
screen "St_Output Bundled_1" 320x240
   IOField "I/O field_9" at 228,67 size 87x20; FormatPattern 999.99
      ProcessValue <- "Data_Real_% label Sloft[1]"
   IOField "I/O field_10" at 228,86 size 87x20; FormatPattern 999.99
      ProcessValue <- "Data_Real_% Unlabel Sloft[1]"
   TextField "Text field_1" at 4,0 size 268x18; Text 'CURRENT SHIFT MINUS 1 ( Output Bundle )'
   IOField "I/O field_2" at 145,86 size 84x20; FormatPattern 9999999
      ProcessValue <- "Data_IntData_Un label Sloft[1]"
   IOField "I/O field_3" at 145,67 size 84x20; FormatPattern 9999999
      ProcessValue <- "Data_IntData_Label Sloft[1]"
   IOField "I/O field_6" at 6,17 size 109x15; FormatPattern 9999999999999999999999999999999999999999
      ProcessValue <- "Data_DTL1_Cur_ShiftA_1"
   TextField "Text field_9" at 120,17 size 18x13; Text 'S/D'
   IOField "I/O field_7" at 143,17 size 109x15; FormatPattern 9999999999999999999999999999999999999999
      ProcessValue <- "Data_DTL1_Cur_ShiftB_1"
   Button "Button_1" at 101,214 size 128x25; TextOff 'Back To Quantity Data'; TextOn 'Page 1'
      on Click: ActivateScreen("St_Quantity Data_1", 0)
   TextField "Text field_5" at 7,86 size 139x20; Text 'Unlabeled Bundle'
   TextField "Text field_4" at 7,67 size 139x20; Text 'Labeled Bundle'
   TextField "Text field_15" at 145,48 size 84x19; Text 'Pcs'
   TextField "Text field_16" at 228,48 size 87x19; Text '% (From input)'
   TextField "Text field_17" at 7,48 size 139x19; Text 'Output Bundle'
   IOField "I/O field_27" at 253,16 size 66x17; FormatPattern ????????
      ProcessValue <- "Data_String_sDT_Machine id"

screen "St_Output Bundled_2" 320x240
   IOField "I/O field_9" at 228,67 size 87x20; FormatPattern 999.99
      ProcessValue <- "Data_Real_% label Sloft[2]"
   IOField "I/O field_10" at 228,86 size 87x20; FormatPattern 999.99
      ProcessValue <- "Data_Real_% Unlabel Sloft[2]"
   TextField "Text field_1" at 4,0 size 262x18; Text 'CURRENT SHIFT MINUS 2 ( Ouput Bundle )'
   IOField "I/O field_2" at 145,86 size 84x20; FormatPattern 9999999
      ProcessValue <- "Data_IntData_Un label Sloft[2]"
   IOField "I/O field_3" at 145,67 size 84x20; FormatPattern 9999999
      ProcessValue <- "Data_IntData_Label Sloft[2]"
   IOField "I/O field_6" at 6,17 size 109x15; FormatPattern 9999999999999999999999999999999999999999
      ProcessValue <- "Data_DTL1_Cur_ShiftA_2"
   TextField "Text field_9" at 120,17 size 18x13; Text 'S/D'
   IOField "I/O field_7" at 143,17 size 109x15; FormatPattern 9999999999999999999999999999999999999999
      ProcessValue <- "Data_DTL1_Cur_ShiftB_2"
   Button "Button_1" at 101,214 size 128x25; TextOff 'Back To Quantity Data'; TextOn 'Page 1'
      on Click: ActivateScreen("St_Quantity Data_2", 0)
   TextField "Text field_5" at 7,86 size 139x20; Text 'Unlabeled Bundle'
   TextField "Text field_4" at 7,67 size 139x20; Text 'Labeled Bundle'
   TextField "Text field_15" at 145,48 size 84x19; Text 'Pcs'
   TextField "Text field_16" at 228,48 size 87x19; Text '% (From input)'
   TextField "Text field_17" at 7,48 size 139x19; Text 'Output Bundle'
   IOField "I/O field_27" at 253,16 size 66x17; FormatPattern ????????
      ProcessValue <- "Data_String_sDT_Machine id"

screen "St_Output Bundled_3" 320x240
   IOField "I/O field_9" at 228,67 size 87x20; FormatPattern 999.99
      ProcessValue <- "Data_Real_% label Sloft[3]"
   IOField "I/O field_10" at 228,86 size 87x20; FormatPattern 999.99
      ProcessValue <- "Data_Real_% Unlabel Sloft[3]"
   TextField "Text field_1" at 4,0 size 268x18; Text 'CURRENT SHIFT MINUS 3 ( Output Bundle )'
   IOField "I/O field_2" at 145,86 size 84x20; FormatPattern 9999999
      ProcessValue <- "Data_IntData_Un label Sloft[3]"
   IOField "I/O field_3" at 145,67 size 84x20; FormatPattern 9999999
      ProcessValue <- "Data_IntData_Label Sloft[3]"
   IOField "I/O field_6" at 6,17 size 109x15; FormatPattern 9999999999999999999999999999999999999999
      ProcessValue <- "Data_DTL1_Cur_ShiftA_3"
   TextField "Text field_9" at 120,17 size 18x13; Text 'S/D'
   IOField "I/O field_7" at 143,17 size 109x15; FormatPattern 9999999999999999999999999999999999999999
      ProcessValue <- "Data_DTL1_Cur_ShiftB_3"
   Button "Button_1" at 101,214 size 128x25; TextOff 'Back To Quantity Data'; TextOn 'Page 1'
      on Click: ActivateScreen("St_Quantity Data_3", 0)
   TextField "Text field_5" at 7,86 size 139x20; Text 'Unlabeled Bundle'
   TextField "Text field_4" at 7,67 size 139x20; Text 'Labeled Bundle'
   TextField "Text field_15" at 145,48 size 84x19; Text 'Pcs'
   TextField "Text field_16" at 228,48 size 87x19; Text '% (From input)'
   TextField "Text field_17" at 7,48 size 139x19; Text 'Output Bundle'
   IOField "I/O field_27" at 253,16 size 66x17; FormatPattern ????????
      ProcessValue <- "Data_String_sDT_Machine id"

screen "St_Output Bundled_4" 320x240
   IOField "I/O field_9" at 228,67 size 87x20; FormatPattern 999.99
      ProcessValue <- "Data_Real_% label Sloft[4]"
   IOField "I/O field_10" at 228,86 size 87x20; FormatPattern 999.99
      ProcessValue <- "Data_Real_% Unlabel Sloft[4]"
   TextField "Text field_1" at 4,0 size 268x18; Text 'CURRENT SHIFT MINUS 4 ( Output Bundle )'
   IOField "I/O field_2" at 145,86 size 84x20; FormatPattern 9999999
      ProcessValue <- "Data_IntData_Un label Sloft[4]"
   IOField "I/O field_3" at 145,67 size 84x20; FormatPattern 9999999
      ProcessValue <- "Data_IntData_Label Sloft[4]"
   TextField "Text field_18" at 230,49 size 14x15; Text '%'
   IOField "I/O field_6" at 6,17 size 109x15; FormatPattern 9999999999999999999999999999999999999999
      ProcessValue <- "Data_DTL1_Cur_ShiftA_4"
   TextField "Text field_9" at 120,17 size 18x13; Text 'S/D'
   IOField "I/O field_7" at 143,17 size 109x15; FormatPattern 9999999999999999999999999999999999999999
      ProcessValue <- "Data_DTL1_Cur_ShiftB_4"
   Button "Button_1" at 101,214 size 128x25; TextOff 'Back To Quantity Data'; TextOn 'Page 1'
      on Click: ActivateScreen("St_Quantity Data_4", 0)
   TextField "Text field_5" at 7,86 size 139x20; Text 'Unlabeled Bundle'
   TextField "Text field_4" at 7,67 size 139x20; Text 'Labeled Bundle'
   TextField "Text field_15" at 145,48 size 84x19; Text 'Pcs'
   TextField "Text field_16" at 228,48 size 87x19; Text '% (From input)'
   TextField "Text field_17" at 7,48 size 139x19; Text 'Output Bundle'
   IOField "I/O field_27" at 253,16 size 66x17; FormatPattern ????????
      ProcessValue <- "Data_String_sDT_Machine id"

screen "St_Output Bundled_5" 320x240
   IOField "I/O field_9" at 228,67 size 87x20; FormatPattern 999.99
      ProcessValue <- "Data_Real_% label Sloft[5]"
   IOField "I/O field_10" at 228,86 size 87x20; FormatPattern 999.99
      ProcessValue <- "Data_Real_% Unlabel Sloft[5]"
   TextField "Text field_5" at 7,86 size 139x20; Text 'Unlabeled Bundle'
   TextField "Text field_1" at 3,0 size 262x18; Text 'CURRENT SHIFT MINUS 5 ( Ouput Bundle )'
   TextField "Text field_4" at 7,67 size 139x20; Text 'Labeled Bundle'
   IOField "I/O field_2" at 145,86 size 84x20; FormatPattern 9999999
      ProcessValue <- "Data_IntData_Un label Sloft[5]"
   IOField "I/O field_3" at 145,67 size 84x20; FormatPattern 9999999
      ProcessValue <- "Data_IntData_Label Sloft[5]"
   TextField "Text field_15" at 145,48 size 84x19; Text 'Pcs'
   TextField "Text field_16" at 228,48 size 87x19; Text '% (From input)'
   TextField "Text field_17" at 7,48 size 139x19; Text 'Output Bundle'
   IOField "I/O field_6" at 6,17 size 109x15; FormatPattern 9999999999999999999999999999999999999999
      ProcessValue <- "Data_DTL1_Cur_ShiftA_5"
   TextField "Text field_9" at 120,17 size 18x13; Text 'S/D'
   IOField "I/O field_7" at 143,17 size 109x15; FormatPattern 9999999999999999999999999999999999999999
      ProcessValue <- "Data_DTL1_Cur_ShiftB_5"
   Button "Button_1" at 101,214 size 128x25; TextOff 'Back To Quantity Data'; TextOn 'Page 1'
      on Click: ActivateScreen("St_Quantity Data_5", 0)
   IOField "I/O field_27" at 253,16 size 66x17; FormatPattern ????????
      ProcessValue <- "Data_String_sDT_Machine id"

screen "St_Quantity Data" 320x240
   Button "Button_4" at 1,78 size 61x38; TextOff 'Labeled Bundle'
      on Click: ActivateScreen("St_Output Bundled", 0)
   Button "Button_5" at 1,114 size 61x55; TextOff 'Unlabeled Bundle'
      on Click: ActivateScreen("St_Output Bundled", 0)
   IOField "I/O field_15" at 232,150 size 87x19; FormatPattern 999.99
      ProcessValue <- "Data_Real_% Sloft bypass[0]"
   IOField "I/O field_16" at 183,150 size 50x19; FormatPattern 9999999
      ProcessValue <- "Data_IntData_Sloft Bypass[0]"
   TextField "Text field_11" at 60,150 size 124x19; Text 'Output - Running Bypass'
   TextField "Text field_8" at 1,41 size 183x19; Text 'Input Bundle'
   IOField "I/O field_13" at 232,132 size 87x19; FormatPattern 999.99
      ProcessValue <- "Data_Real_%Bad Read[0]"
   IOField "I/O field_12" at 183,132 size 50x19; FormatPattern 9999999
      ProcessValue <- "Data_IntData_Bad R"
   TextField "Text field_6" at 60,132 size 124x19; Text 'Reject Bad Read'
   IOField "I/O field_11" at 232,168 size 87x19; FormatPattern 999.99
      ProcessValue <- "Data_Real_% Total Output[0]"
   IOField "I/O field_9" at 232,78 size 87x19; FormatPattern 999.99
      ProcessValue <- "Data_Real_%Good Read[0]"
   IOField "I/O field_10" at 232,96 size 87x19; FormatPattern 999.99
      ProcessValue <- "Data_Real_% Reject Out Stop[0]"
   IOField "I/O field_8" at 232,114 size 87x19; FormatPattern 999.99
      ProcessValue <- "Data_Real_%InputReject[0]"
   TextField "Text field_5" at 60,96 size 124x19; Text 'Downstream Jammed Reject'
   TextField "Text field_1" at 3,0 size 211x18; Text 'CURRENT SHIFT ( Quantity data )'
   IOField "I/O field_1" at 183,41 size 87x19; FormatPattern 9999999999; Unit  Pcs
      ProcessValue <- "Data_IntData_Input Sloft"
   TextField "Text field_3" at 1,168 size 183x19; Text 'Total Output Bundle'
   TextField "Text field_4" at 60,78 size 124x19; Text 'Output Good Read'
   TextField "Text field_7" at 60,114 size 124x19; Text 'Input Chute Reject'
   IOField "I/O field_2" at 183,96 size 50x19; FormatPattern 9999999
      ProcessValue <- "Data_IntData_Reject Out S"
   IOField "I/O field_3" at 183,78 size 50x19; FormatPattern 9999999
      ProcessValue <- "Data_IntData_Good R"
   IOField "I/O field_5" at 183,168 size 50x19; FormatPattern 9999999
      ProcessValue <- "Data_IntData_Tot Out Slof"
   IOField "I/O field_4" at 183,114 size 50x19; FormatPattern 9999999
      ProcessValue <- "Data_IntData_InReject"
   TextField "Text field_2" at 260,0 size 57x15; Text 'Page 1 of 3'
   Button "Button_1" at 46,213 size 90x25; TextOff 'Statistic Data'
      on Click: ActivateScreen("St_Data Statistic", 0)
   Button "Button_3" at 1,213 size 41x25; TextOff 'Main Page'; PictureOff "Home"
      on Click: ActivateScreen("Main Page", 0)
   Button "Button_2" at 237,213 size 80x25; TextOff 'Next Page -->'; TextOn 'Page 2'
      on Click: ActivateScreen("St_Time machine data", 0)
   TextField "Text field_10" at 1,189 size 184x20; Text 'Applicator Freeze'
   IOField "I/O field_14" at 182,189 size 87x20; FormatPattern 999; Unit   Times
      ProcessValue <- "Data_IntData_uintDT_AplicatorFreeze[0]"
   TextField "Text field_15" at 183,60 size 50x19; Text 'Pcs'
   TextField "Text field_16" at 232,60 size 87x19; Text '% (From Input )'
   TextField "Text field_17" at 1,60 size 183x19; Text 'Detail Output Bundle'
   IOField "I/O field_6" at 6,17 size 109x15; FormatPattern 9999999999999999999999999999999999999999
      ProcessValue <- "Data_DTL1_Cur_ShiftA"
   TextField "Text field_9" at 120,17 size 18x13; Text 'S/D'
   IOField "I/O field_7" at 143,17 size 109x15; FormatPattern 9999999999999999999999999999999999999999
      ProcessValue <- "Data_DTL1_Cur_ShiftB"
   IOField "I/O field_27" at 253,16 size 66x17; FormatPattern ????????
      ProcessValue <- "Data_String_sDT_Machine id"

screen "St_Quantity Data_1" 320x240
   Button "Button_4" at 1,78 size 61x38; TextOff 'Labeled Bundled'
      on Click: ActivateScreen("St_Output Bundled_1", 0)
   Button "Button_5" at 1,114 size 61x55; TextOff 'Unlabeled Bundled'
      on Click: ActivateScreen("St_Output Bundled_1", 0)
   IOField "I/O field_15" at 232,150 size 87x19; FormatPattern 999.99
      ProcessValue <- "Data_Real_% Sloft bypass[1]"
   IOField "I/O field_16" at 183,150 size 50x19; FormatPattern 9999999
      ProcessValue <- "Data_IntData_Sloft Bypass[1]"
   TextField "Text field_11" at 60,150 size 124x19; Text 'Output - Running Bypass'
   TextField "Text field_8" at 1,41 size 183x19; Text 'Input Bundle'
   IOField "I/O field_13" at 232,132 size 87x19; FormatPattern 999.99
      ProcessValue <- "Data_Real_%Bad Read[1]"
   IOField "I/O field_12" at 183,132 size 50x19; FormatPattern 9999999
      ProcessValue <- "Data_IntData_Bad R_1"
   TextField "Text field_6" at 60,132 size 124x19; Text 'Reject Bad Read'
   IOField "I/O field_11" at 232,168 size 87x19; FormatPattern 999.99
      ProcessValue <- "Data_Real_% Total Output[1]"
   IOField "I/O field_9" at 232,78 size 87x19; FormatPattern 999.99
      ProcessValue <- "Data_Real_%Good Read[1]"
   IOField "I/O field_10" at 232,96 size 87x19; FormatPattern 999.99
      ProcessValue <- "Data_Real_% Reject Out Stop[1]"
   IOField "I/O field_8" at 232,114 size 87x19; FormatPattern 999.99
      ProcessValue <- "Data_Real_%InputReject[1]"
   TextField "Text field_5" at 60,96 size 124x19; Text 'Downstream Jammed Reject'
   TextField "Text field_1" at 3,0 size 155x18; Text 'CURRENT SHIFT MINUS 1'
   IOField "I/O field_1" at 183,41 size 87x19; FormatPattern 9999999999; Unit  Pcs
      ProcessValue <- "Data_IntData_Input Sloft_1"
   TextField "Text field_3" at 1,168 size 183x19; Text 'Total Output Bundle'
   TextField "Text field_4" at 60,78 size 124x19; Text 'Output Good Read'
   TextField "Text field_7" at 60,114 size 124x19; Text 'Input Chute Reject'
   IOField "I/O field_2" at 183,96 size 50x19; FormatPattern 9999999
      ProcessValue <- "Data_IntData_Reject Out S_1"
   IOField "I/O field_3" at 183,78 size 50x19; FormatPattern 9999999
      ProcessValue <- "Data_IntData_Good R_1"
   IOField "I/O field_5" at 183,168 size 50x19; FormatPattern 9999999
      ProcessValue <- "Data_IntData_Tot Out Slof_1"
   IOField "I/O field_4" at 183,114 size 50x19; FormatPattern 9999999
      ProcessValue <- "Data_IntData_InReject_1"
   TextField "Text field_2" at 260,0 size 57x15; Text 'Page 1 of 3'
   Button "Button_1" at 46,213 size 90x25; TextOff 'Statistic Data'
      on Click: ActivateScreen("St_Data Statistic", 0)
   Button "Button_3" at 1,213 size 41x25; TextOff 'Main Page'; PictureOff "Home"
      on Click: ActivateScreen("Main Page", 0)
   Button "Button_2" at 237,213 size 80x25; TextOff 'Next Page -->'; TextOn 'Page 2'
      on Click: ActivateScreen("St_Time machine data_1", 0)
   TextField "Text field_10" at 1,189 size 184x20; Text 'Applicator Freeze'
   IOField "I/O field_14" at 182,189 size 87x20; FormatPattern 999; Unit   Times
      ProcessValue <- "Data_IntData_uintDT_AplicatorFreeze[1]"
   IOField "I/O field_6" at 6,17 size 109x15; FormatPattern 9999999999999999999999999999999999999999
      ProcessValue <- "Data_DTL1_Cur_ShiftA_1"
   TextField "Text field_9" at 120,17 size 18x13; Text 'S/D'
   IOField "I/O field_7" at 143,17 size 109x15; FormatPattern 9999999999999999999999999999999999999999
      ProcessValue <- "Data_DTL1_Cur_ShiftB_1"
   TextField "Text field_15" at 183,60 size 50x19; Text 'Pcs'
   TextField "Text field_16" at 232,60 size 87x19; Text '% (From Input )'
   TextField "Text field_17" at 1,60 size 183x19; Text 'Detail Output Bundle'
   IOField "I/O field_27" at 253,16 size 66x17; FormatPattern ????????
      ProcessValue <- "Data_String_sDT_Machine id"

screen "St_Quantity Data_2" 320x240
   Button "Button_4" at 1,78 size 61x37; TextOff 'Labeled Bundle'
      on Click: ActivateScreen("St_Output Bundled_2", 0)
   Button "Button_5" at 1,114 size 61x56; TextOff 'Unlabeled Bundle'
      on Click: ActivateScreen("St_Output Bundled_2", 0)
   IOField "I/O field_15" at 232,150 size 87x19; FormatPattern 999.99
      ProcessValue <- "Data_Real_% Sloft bypass[2]"
   IOField "I/O field_16" at 183,150 size 50x19; FormatPattern 9999999
      ProcessValue <- "Data_IntData_Sloft Bypass[2]"
   TextField "Text field_11" at 60,150 size 124x19; Text 'Output - Running Bypass'
   TextField "Text field_8" at 1,41 size 183x19; Text 'Input Bundle'
   IOField "I/O field_13" at 232,132 size 87x19; FormatPattern 999.99
      ProcessValue <- "Data_Real_%Bad Read[2]"
   IOField "I/O field_12" at 183,132 size 50x19; FormatPattern 9999999
      ProcessValue <- "Data_IntData_Bad R_2"
   TextField "Text field_6" at 60,132 size 124x19; Text 'Reject Bad Read'
   IOField "I/O field_11" at 232,168 size 87x19; FormatPattern 999.99
      ProcessValue <- "Data_Real_% Total Output[2]"
   IOField "I/O field_9" at 232,78 size 87x19; FormatPattern 999.99
      ProcessValue <- "Data_Real_%Good Read[2]"
   IOField "I/O field_10" at 232,96 size 87x19; FormatPattern 999.99
      ProcessValue <- "Data_Real_% Reject Out Stop[2]"
   IOField "I/O field_8" at 232,114 size 87x19; FormatPattern 999.99
      ProcessValue <- "Data_Real_%InputReject[2]"
   TextField "Text field_5" at 60,96 size 124x19; Text 'Downstream Jammed Reject'
   TextField "Text field_1" at 3,0 size 155x18; Text 'CURRENT SHIFT MINUS 2'
   IOField "I/O field_1" at 183,41 size 87x19; FormatPattern 9999999999; Unit  Pcs
      ProcessValue <- "Data_IntData_Input Sloft_2"
   TextField "Text field_3" at 1,168 size 183x19; Text 'Total Output Bundle'
   TextField "Text field_4" at 60,78 size 124x19; Text 'Output Good Read'
   TextField "Text field_7" at 60,114 size 124x19; Text 'Input Chute Reject'
   IOField "I/O field_2" at 183,96 size 50x19; FormatPattern 9999999
      ProcessValue <- "Data_IntData_Reject Out S_2"
   IOField "I/O field_3" at 183,78 size 50x19; FormatPattern 9999999
      ProcessValue <- "Data_IntData_Good R_2"
   IOField "I/O field_5" at 183,168 size 50x19; FormatPattern 9999999
      ProcessValue <- "Data_IntData_Tot Out Slof_2"
   IOField "I/O field_4" at 183,114 size 50x19; FormatPattern 9999999
      ProcessValue <- "Data_IntData_InReject_2"
   TextField "Text field_2" at 260,0 size 57x15; Text 'Page 1 of 3'
   Button "Button_1" at 46,213 size 90x25; TextOff 'Statistic Data'
      on Click: ActivateScreen("St_Data Statistic", 0)
   Button "Button_3" at 1,213 size 41x25; TextOff 'Main Page'; PictureOff "Home"
      on Click: ActivateScreen("Main Page", 0)
   Button "Button_2" at 237,213 size 80x25; TextOff 'Next Page -->'; TextOn 'Page 2'
      on Click: ActivateScreen("St_Time machine data_2", 0)
   TextField "Text field_10" at 1,189 size 184x20; Text 'Applicator Freeze'
   IOField "I/O field_14" at 182,189 size 87x20; FormatPattern 999; Unit   Times
      ProcessValue <- "Data_IntData_uintDT_AplicatorFreeze[2]"
   IOField "I/O field_6" at 6,17 size 109x15; FormatPattern 9999999999999999999999999999999999999999
      ProcessValue <- "Data_DTL1_Cur_ShiftA_2"
   TextField "Text field_9" at 120,17 size 18x13; Text 'S/D'
   IOField "I/O field_7" at 143,17 size 109x15; FormatPattern 9999999999999999999999999999999999999999
      ProcessValue <- "Data_DTL1_Cur_ShiftB_2"
   TextField "Text field_15" at 183,60 size 50x19; Text 'Pcs'
   TextField "Text field_16" at 232,60 size 87x19; Text '% (From Input )'
   TextField "Text field_17" at 1,60 size 183x19; Text 'Detail Output Bundle'
   IOField "I/O field_27" at 253,16 size 66x17; FormatPattern ????????
      ProcessValue <- "Data_String_sDT_Machine id"

screen "St_Quantity Data_3" 320x240
   Button "Button_4" at 1,78 size 61x38; TextOff 'Labeled Bundle'
      on Click: ActivateScreen("St_Output Bundled_3", 0)
   Button "Button_5" at 1,114 size 61x57; TextOff 'Unlabeled Bundle'
      on Click: ActivateScreen("St_Output Bundled_3", 0)
   IOField "I/O field_15" at 232,150 size 87x19; FormatPattern 999.99
      ProcessValue <- "Data_Real_% Sloft bypass[3]"
   IOField "I/O field_16" at 183,150 size 50x19; FormatPattern 9999999
      ProcessValue <- "Data_IntData_Sloft Bypass[3]"
   TextField "Text field_11" at 60,150 size 124x19; Text 'Output - Running Bypass'
   TextField "Text field_8" at 1,41 size 183x19; Text 'Input Bundle'
   IOField "I/O field_13" at 232,132 size 87x19; FormatPattern 999.99
      ProcessValue <- "Data_Real_%Bad Read[3]"
   IOField "I/O field_12" at 183,132 size 50x19; FormatPattern 9999999
      ProcessValue <- "Data_IntData_Bad R_3"
   TextField "Text field_6" at 60,132 size 124x19; Text 'Reject Bad Read'
   IOField "I/O field_11" at 232,168 size 87x19; FormatPattern 999.99
      ProcessValue <- "Data_Real_% Total Output[3]"
   IOField "I/O field_9" at 232,78 size 87x19; FormatPattern 999.99
      ProcessValue <- "Data_Real_%Good Read[3]"
   IOField "I/O field_10" at 232,96 size 87x19; FormatPattern 999.99
      ProcessValue <- "Data_Real_% Reject Out Stop[3]"
   IOField "I/O field_8" at 232,114 size 87x19; FormatPattern 999.99
      ProcessValue <- "Data_Real_%InputReject[3]"
   TextField "Text field_5" at 60,96 size 124x19; Text 'Downstream Jammed Reject'
   TextField "Text field_1" at 3,0 size 155x18; Text 'CURRENT SHIFT MINUS 3'
   IOField "I/O field_1" at 183,41 size 87x19; FormatPattern 9999999999; Unit  Pcs
      ProcessValue <- "Data_IntData_Input Sloft_3"
   TextField "Text field_3" at 1,168 size 183x19; Text 'Total Output Bundle'
   TextField "Text field_4" at 60,78 size 124x19; Text 'Output Good Read'
   TextField "Text field_7" at 60,114 size 124x19; Text 'Input Chute Reject'
   IOField "I/O field_2" at 183,96 size 50x19; FormatPattern 9999999
      ProcessValue <- "Data_IntData_Reject Out S_3"
   IOField "I/O field_3" at 183,78 size 50x19; FormatPattern 9999999
      ProcessValue <- "Data_IntData_Good R_3"
   IOField "I/O field_5" at 183,168 size 50x19; FormatPattern 9999999
      ProcessValue <- "Data_IntData_Tot Out Slof_3"
   IOField "I/O field_4" at 183,114 size 50x19; FormatPattern 9999999
      ProcessValue <- "Data_IntData_InReject_3"
   TextField "Text field_2" at 260,0 size 57x15; Text 'Page 1 of 3'
   Button "Button_1" at 46,213 size 90x25; TextOff 'Statistic Data'
      on Click: ActivateScreen("St_Data Statistic", 0)
   Button "Button_3" at 1,213 size 41x25; TextOff 'Main Page'; PictureOff "Home"
      on Click: ActivateScreen("Main Page", 0)
   Button "Button_2" at 237,213 size 80x25; TextOff 'Next Page -->'; TextOn 'Page 2'
      on Click: ActivateScreen("St_Time machine data_3", 0)
   TextField "Text field_10" at 1,189 size 184x20; Text 'Applicator Freeze'
   IOField "I/O field_14" at 182,189 size 87x20; FormatPattern 999; Unit   Times
      ProcessValue <- "Data_IntData_uintDT_AplicatorFreeze[3]"
   IOField "I/O field_6" at 6,17 size 109x15; FormatPattern 9999999999999999999999999999999999999999
      ProcessValue <- "Data_DTL1_Cur_ShiftA_3"
   TextField "Text field_9" at 120,17 size 18x13; Text 'S/D'
   IOField "I/O field_7" at 143,17 size 109x15; FormatPattern 9999999999999999999999999999999999999999
      ProcessValue <- "Data_DTL1_Cur_ShiftB_3"
   TextField "Text field_15" at 183,60 size 50x19; Text 'Pcs'
   TextField "Text field_16" at 232,60 size 87x19; Text '% (From Input )'
   TextField "Text field_17" at 1,60 size 183x19; Text 'Detail Output Bundle'
   IOField "I/O field_27" at 253,16 size 66x17; FormatPattern ????????
      ProcessValue <- "Data_String_sDT_Machine id"

screen "St_Quantity Data_4" 320x240
   Button "Button_4" at 1,78 size 61x38; TextOff 'Labeled Bundle'
      on Click: ActivateScreen("St_Output Bundled_4", 0)
   Button "Button_5" at 1,114 size 61x57; TextOff 'Unlabeled Bundle'
      on Click: ActivateScreen("St_Output Bundled_4", 0)
   IOField "I/O field_15" at 232,150 size 87x19; FormatPattern 999.99
      ProcessValue <- "Data_Real_% Sloft bypass[4]"
   IOField "I/O field_16" at 183,150 size 50x19; FormatPattern 9999999
      ProcessValue <- "Data_IntData_Sloft Bypass[4]"
   TextField "Text field_11" at 60,150 size 124x19; Text 'Output - Running Bypass'
   TextField "Text field_8" at 1,41 size 183x19; Text 'Input Bundle'
   IOField "I/O field_13" at 232,132 size 87x19; FormatPattern 999.99
      ProcessValue <- "Data_Real_%Bad Read[4]"
   IOField "I/O field_12" at 183,132 size 50x19; FormatPattern 9999999
      ProcessValue <- "Data_IntData_Bad R_4"
   TextField "Text field_6" at 60,132 size 124x19; Text 'Reject Bad Read'
   IOField "I/O field_11" at 232,168 size 87x19; FormatPattern 999.99
      ProcessValue <- "Data_Real_% Total Output[4]"
   IOField "I/O field_9" at 232,78 size 87x19; FormatPattern 999.99
      ProcessValue <- "Data_Real_%Good Read[4]"
   IOField "I/O field_10" at 232,96 size 87x19; FormatPattern 999.99
      ProcessValue <- "Data_Real_% Reject Out Stop[4]"
   IOField "I/O field_8" at 232,114 size 87x19; FormatPattern 999.99
      ProcessValue <- "Data_Real_%InputReject[4]"
   TextField "Text field_5" at 60,96 size 124x19; Text 'Downstream Jammed Reject'
   TextField "Text field_1" at 3,0 size 155x18; Text 'CURRENT SHIFT MINUS 4'
   IOField "I/O field_1" at 183,41 size 87x19; FormatPattern 9999999999; Unit  Pcs
      ProcessValue <- "Data_IntData_Input Sloft_4"
   TextField "Text field_3" at 1,168 size 183x19; Text 'Total Output Bundle'
   TextField "Text field_4" at 60,78 size 124x19; Text 'Output Good Read'
   TextField "Text field_7" at 60,114 size 124x19; Text 'Input Chute Reject'
   IOField "I/O field_2" at 183,96 size 50x19; FormatPattern 9999999
      ProcessValue <- "Data_IntData_Reject Out S_4"
   IOField "I/O field_3" at 183,78 size 50x19; FormatPattern 9999999
      ProcessValue <- "Data_IntData_Good R_4"
   IOField "I/O field_5" at 183,168 size 50x19; FormatPattern 9999999
      ProcessValue <- "Data_IntData_Tot Out Slof_4"
   IOField "I/O field_4" at 183,114 size 50x19; FormatPattern 9999999
      ProcessValue <- "Data_IntData_InReject_4"
   TextField "Text field_2" at 260,0 size 57x15; Text 'Page 1 of 3'
   Button "Button_1" at 46,213 size 90x25; TextOff 'Statistic Data'
      on Click: ActivateScreen("St_Data Statistic", 0)
   Button "Button_3" at 1,213 size 41x25; TextOff 'Main Page'; PictureOff "Home"
      on Click: ActivateScreen("Main Page", 0)
   Button "Button_2" at 237,213 size 80x25; TextOff 'Next Page -->'; TextOn 'Page 2'
      on Click: ActivateScreen("St_Time machine data_4", 0)
   TextField "Text field_10" at 1,189 size 184x20; Text 'Applicator Freeze'
   IOField "I/O field_14" at 182,189 size 87x20; FormatPattern 999; Unit   Times
      ProcessValue <- "Data_IntData_uintDT_AplicatorFreeze[4]"
   IOField "I/O field_6" at 6,17 size 109x15; FormatPattern 9999999999999999999999999999999999999999
      ProcessValue <- "Data_DTL1_Cur_ShiftA_4"
   TextField "Text field_9" at 120,17 size 18x13; Text 'S/D'
   IOField "I/O field_7" at 143,17 size 109x15; FormatPattern 9999999999999999999999999999999999999999
      ProcessValue <- "Data_DTL1_Cur_ShiftB_4"
   TextField "Text field_15" at 183,60 size 50x19; Text 'Pcs'
   TextField "Text field_16" at 232,60 size 87x19; Text '% (From Input )'
   TextField "Text field_17" at 1,60 size 183x19; Text 'Detail Output Bundle'
   IOField "I/O field_27" at 253,16 size 66x17; FormatPattern ????????
      ProcessValue <- "Data_String_sDT_Machine id"

screen "St_Quantity Data_5" 320x240
   Button "Button_4" at 1,78 size 61x38; TextOff 'Labeled Bundle'
      on Click: ActivateScreen("St_Output Bundled_5", 0)
   Button "Button_5" at 1,114 size 61x57; TextOff 'Unlabeled Bundle'
      on Click: ActivateScreen("St_Output Bundled_5", 0)
   IOField "I/O field_15" at 232,150 size 87x19; FormatPattern 999.99
      ProcessValue <- "Data_Real_% Sloft bypass[5]"
   IOField "I/O field_16" at 183,150 size 50x19; FormatPattern 9999999
      ProcessValue <- "Data_IntData_Sloft Bypass[5]"
   TextField "Text field_11" at 60,150 size 124x19; Text 'Output - Running Bypass'
   TextField "Text field_8" at 1,41 size 183x19; Text 'Input Bundle'
   IOField "I/O field_13" at 232,132 size 87x19; FormatPattern 999.99
      ProcessValue <- "Data_Real_%Bad Read[5]"
   IOField "I/O field_12" at 183,132 size 50x19; FormatPattern 9999999
      ProcessValue <- "Data_IntData_Bad R_5"
   TextField "Text field_6" at 60,132 size 124x19; Text 'Reject Bad Read'
   IOField "I/O field_11" at 232,168 size 87x19; FormatPattern 999.99
      ProcessValue <- "Data_Real_% Total Output[5]"
   IOField "I/O field_9" at 232,78 size 87x19; FormatPattern 999.99
      ProcessValue <- "Data_Real_%Good Read[5]"
   IOField "I/O field_10" at 232,96 size 87x19; FormatPattern 999.99
      ProcessValue <- "Data_Real_% Reject Out Stop[5]"
   IOField "I/O field_8" at 232,114 size 87x19; FormatPattern 999.99
      ProcessValue <- "Data_Real_%InputReject[5]"
   TextField "Text field_5" at 60,96 size 124x19; Text 'Downstream Jammed Reject'
   TextField "Text field_1" at 3,0 size 155x18; Text 'CURRENT SHIFT MINUS 5'
   IOField "I/O field_1" at 183,41 size 87x19; FormatPattern 9999999999; Unit  Pcs
      ProcessValue <- "Data_IntData_Input Sloft_5"
   TextField "Text field_3" at 1,168 size 183x19; Text 'Total Output Bundle'
   TextField "Text field_4" at 60,78 size 124x19; Text 'Output Good Read'
   TextField "Text field_7" at 60,114 size 124x19; Text 'Input Chute Reject'
   IOField "I/O field_2" at 183,96 size 50x19; FormatPattern 9999999
      ProcessValue <- "Data_IntData_Reject Out S_5"
   IOField "I/O field_3" at 183,78 size 50x19; FormatPattern 9999999
      ProcessValue <- "Data_IntData_Good R_5"
   IOField "I/O field_5" at 183,168 size 50x19; FormatPattern 9999999
      ProcessValue <- "Data_IntData_Tot Out Slof_5"
   IOField "I/O field_4" at 183,114 size 50x19; FormatPattern 9999999
      ProcessValue <- "Data_IntData_InReject_5"
   TextField "Text field_2" at 260,0 size 57x15; Text 'Page 1 of 3'
   Button "Button_1" at 46,213 size 90x25; TextOff 'Statistic Data'
      on Click: ActivateScreen("St_Data Statistic", 0)
   Button "Button_3" at 1,213 size 41x25; TextOff 'Main Page'; PictureOff "Home"
      on Click: ActivateScreen("Main Page", 0)
   Button "Button_2" at 237,213 size 80x25; TextOff 'Next Page -->'; TextOn 'Page 2'
      on Click: ActivateScreen("St_Time machine data_5", 0)
   TextField "Text field_10" at 1,189 size 184x20; Text 'Applicator Freeze'
   IOField "I/O field_14" at 182,189 size 87x20; FormatPattern 999; Unit   Times
      ProcessValue <- "Data_IntData_uintDT_AplicatorFreeze[5]"
   IOField "I/O field_6" at 6,17 size 109x15; FormatPattern 9999999999999999999999999999999999999999
      ProcessValue <- "Data_DTL1_Cur_ShiftA_5"
   TextField "Text field_9" at 120,17 size 18x13; Text 'S/D'
   IOField "I/O field_7" at 143,17 size 109x15; FormatPattern 9999999999999999999999999999999999999999
      ProcessValue <- "Data_DTL1_Cur_ShiftB_5"
   TextField "Text field_15" at 183,60 size 50x19; Text 'Pcs'
   TextField "Text field_16" at 232,60 size 87x19; Text '% (From Input )'
   TextField "Text field_17" at 1,60 size 183x19; Text 'Detail Output Bundle'
   IOField "I/O field_27" at 253,16 size 66x17; FormatPattern ????????
      ProcessValue <- "Data_String_sDT_Machine id"

screen "St_Time machine data" 320x240
   IOField "I/O field_13" at 243,83 size 56x19; FormatPattern 999.99; Unit   %
      ProcessValue <- "Data_Real_%Mesin Stop[0]"
   IOField "I/O field_14" at 243,101 size 56x19; FormatPattern 999.99; Unit   %
      ProcessValue <- "Data_Real_%Mesin Run Baypass[0]"
   IOField "I/O field_11" at 243,66 size 56x19; FormatPattern 999.99; Unit   %
      ProcessValue <- "Data_Real_%Mesin Run[0]"
   Button "Button_1" at 46,213 size 90x25; TextOff 'Statistic Data'
      on Click: ActivateScreen("St_Data Statistic", 0)
   Button "Button_3" at 1,213 size 41x25; TextOff 'Main Page'; PictureOff "Home"
      on Click: ActivateScreen("Main Page", 0)
   Button "Button_2" at 237,213 size 80x25; TextOff 'Next page -->'; TextOn 'Page 3'
      on Click: ActivateScreen("St_Error Counter", 0)
   TextField "Text field_1" at 3,0 size 227x18; Text 'CURRENT SHIFT (Time machine data)'
   TextField "Text field_31" at 7,101 size 21x19; Text '3'
   TextField "Text field_30" at 7,83 size 21x19; Text '2'
   TextField "Text field_29" at 7,66 size 21x19; Text '1'
   TextField "Text field_28" at 7,48 size 21x19; Text 'No'
   IOField "I/O field_21" at 219,83 size 25x19; FormatPattern 999
      ProcessValue <- "Data_DTLData_DTL_Mesin Stop[0].SECOND"
   IOField "I/O field_22" at 195,83 size 25x19; FormatPattern 999
      ProcessValue <- "Data_DTLData_DTL_Mesin Stop[0].MINUTE"
   IOField "I/O field_23" at 171,84 size 25x19; FormatPattern 999
      ProcessValue <- "Data_DTLData_DTL_Mesin Stop[0].HOUR"
   TextField "Text field_25" at 27,83 size 145x19; Text 'Stop'
   IOField "I/O field_4" at 219,101 size 25x19; FormatPattern 999
      ProcessValue <- "Data_DTLData_DTL_Mesin Run Baypass[0].SECOND"
   IOField "I/O field_5" at 195,101 size 25x19; FormatPattern 999
      ProcessValue <- "Data_DTLData_DTL_Mesin Run Baypass[0].MINUTE"
   IOField "I/O field_9" at 171,101 size 25x19; FormatPattern 999
      ProcessValue <- "Data_DTLData_DTL_Mesin Run Baypass[0].HOUR"
   TextField "Text field_12" at 219,48 size 25x19; Text 'Sec'
   TextField "Text field_11" at 195,48 size 25x19; Text 'Min'
   IOField "I/O field_2" at 219,66 size 25x19; FormatPattern 999
      ProcessValue <- "Data_DTLData_DTL_Mesin Run[0].SECOND"
   IOField "I/O field_3" at 195,66 size 25x19; FormatPattern 999
      ProcessValue <- "Data_DTLData_DTL_Mesin Run[0].MINUTE"
   TextField "Text field_3" at 27,48 size 145x19; Text 'Time Counter Machine'
   TextField "Text field_4" at 27,66 size 145x19; Text 'Running'
   TextField "Text field_5" at 27,101 size 145x19; Text 'Running Bypass'
   IOField "I/O field_24" at 171,66 size 25x19; FormatPattern 999
      ProcessValue <- "Data_DTLData_DTL_Mesin Run[0].HOUR"
   Button "Button_4" at 151,213 size 80x25; TextOff '<-- Back Page'; TextOn 'Page 1'
      on Click: ActivateScreen("St_Quantity Data", 0)
   TextField "Text field_6" at 260,0 size 57x15; Text 'Page 2 of 3'
   IOField "I/O field_1" at 243,119 size 56x19; FormatPattern 999.99; Unit   %
      ProcessValue <- "Data_Real_%Mesin Error[0]"
   TextField "Text field_7" at 7,119 size 21x19; Text '4'
   IOField "I/O field_8" at 219,119 size 25x19; FormatPattern 999
      ProcessValue <- "Data_DTLData_DTL_Mesin Error[0].SECOND"
   IOField "I/O field_10" at 195,119 size 25x19; FormatPattern 999
      ProcessValue <- "Data_DTLData_DTL_Mesin Error[0].MINUTE"
   IOField "I/O field_12" at 171,119 size 25x19; FormatPattern 999
      ProcessValue <- "Data_DTLData_DTL_Mesin Error[0].HOUR"
   TextField "Text field_8" at 27,119 size 145x19; Text 'Error'
   TextField "Text field_2" at 171,48 size 25x19; Text 'Hour'
   IOField "I/O field_6" at 6,17 size 109x15; FormatPattern 9999999999999999999999999999999999999999
      ProcessValue <- "Data_DTL1_Cur_ShiftA"
   TextField "Text field_9" at 120,17 size 18x13; Text 'S/D'
   IOField "I/O field_7" at 143,17 size 109x15; FormatPattern 9999999999999999999999999999999999999999
      ProcessValue <- "Data_DTL1_Cur_ShiftB"
   IOField "I/O field_16" at 219,138 size 25x19; FormatPattern 999
      ProcessValue <- "Data_DTLData_Total Time Machine[0].SECOND"
   IOField "I/O field_17" at 195,138 size 25x19; FormatPattern 999
      ProcessValue <- "Data_DTLData_Total Time Machine[0].MINUTE"
   IOField "I/O field_18" at 171,138 size 25x19; FormatPattern 999
      ProcessValue <- "Data_DTLData_Total Time Machine[0].HOUR"
   TextField "Text field_10" at 27,138 size 145x19; Text 'Total'
   IOField "I/O field_27" at 253,16 size 66x17; FormatPattern ????????
      ProcessValue <- "Data_String_sDT_Machine id"
   Softkey "Softkey_F1" at 1,202 size 53x38
      on KeyDown: ActivateScreen("Main Page", 0)

screen "St_Time machine data_1" 320x240
   IOField "I/O field_13" at 243,83 size 56x19; FormatPattern 999.99; Unit   %
      ProcessValue <- "Data_Real_%Mesin Stop[1]"
   IOField "I/O field_14" at 243,101 size 56x19; FormatPattern 999.99; Unit   %
      ProcessValue <- "Data_Real_%Mesin Run Baypass[1]"
   IOField "I/O field_11" at 243,66 size 56x19; FormatPattern 999.99; Unit   %
      ProcessValue <- "Data_Real_%Mesin Run[1]"
   Button "Button_1" at 46,213 size 90x25; TextOff 'Statistic Data'
      on Click: ActivateScreen("St_Data Statistic", 0)
   Button "Button_3" at 1,213 size 41x25; TextOff 'Main Page'; PictureOff "Home"
      on Click: ActivateScreen("Main Page", 0)
   Button "Button_2" at 237,213 size 80x25; TextOff 'Next page -->'; TextOn 'Page 3'
      on Click: ActivateScreen("ST_Error Counter_1", 0)
   TextField "Text field_1" at 3,0 size 155x18; Text 'CURRENT SHIFT MINUS 1'
   TextField "Text field_31" at 7,101 size 21x19; Text '3'
   TextField "Text field_30" at 7,83 size 21x19; Text '2'
   TextField "Text field_29" at 7,66 size 21x19; Text '1'
   TextField "Text field_28" at 7,48 size 21x19; Text 'No'
   IOField "I/O field_21" at 219,83 size 25x19; FormatPattern 999
      ProcessValue <- "Data_DTLData_DTL_Mesin Stop[1].SECOND"
   IOField "I/O field_22" at 195,83 size 25x19; FormatPattern 999
      ProcessValue <- "Data_DTLData_DTL_Mesin Stop[1].MINUTE"
   IOField "I/O field_23" at 171,84 size 25x19; FormatPattern 999
      ProcessValue <- "Data_DTLData_DTL_Mesin Stop[1].HOUR"
   TextField "Text field_25" at 27,83 size 145x19; Text 'Stop'
   IOField "I/O field_4" at 219,101 size 25x19; FormatPattern 999
      ProcessValue <- "Data_DTLData_DTL_Mesin Run Baypass[1].SECOND"
   IOField "I/O field_5" at 195,101 size 25x19; FormatPattern 999
      ProcessValue <- "Data_DTLData_DTL_Mesin Run Baypass[1].MINUTE"
   IOField "I/O field_9" at 171,101 size 25x19; FormatPattern 999
      ProcessValue <- "Data_DTLData_DTL_Mesin Run Baypass[1].HOUR"
   TextField "Text field_12" at 219,48 size 25x19; Text 'Sec'
   TextField "Text field_11" at 195,48 size 25x19; Text 'Min'
   IOField "I/O field_2" at 219,66 size 25x19; FormatPattern 999
      ProcessValue <- "Data_DTLData_DTL_Mesin Run[1].SECOND"
   IOField "I/O field_3" at 195,66 size 25x19; FormatPattern 999
      ProcessValue <- "Data_DTLData_DTL_Mesin Run[1].MINUTE"
   TextField "Text field_3" at 27,48 size 145x19; Text 'Time Counter Machine'
   TextField "Text field_4" at 27,66 size 145x19; Text 'Running'
   TextField "Text field_5" at 27,101 size 145x19; Text 'Running Bypass'
   IOField "I/O field_24" at 171,66 size 25x19; FormatPattern 999
      ProcessValue <- "Data_DTLData_DTL_Mesin Run[1].HOUR"
   Button "Button_4" at 151,213 size 80x25; TextOff '<-- Back Page'; TextOn 'Page 1'
      on Click: ActivateScreen("St_Quantity Data_1", 0)
   TextField "Text field_6" at 260,0 size 57x15; Text 'Page 2 of 3'
   IOField "I/O field_1" at 243,119 size 56x19; FormatPattern 999.99; Unit   %
      ProcessValue <- "Data_Real_%Mesin Error[1]"
   TextField "Text field_7" at 7,119 size 21x19; Text '4'
   IOField "I/O field_8" at 219,119 size 25x19; FormatPattern 999
      ProcessValue <- "Data_DTLData_DTL_Mesin Error[1].SECOND"
   IOField "I/O field_10" at 195,119 size 25x19; FormatPattern 999
      ProcessValue <- "Data_DTLData_DTL_Mesin Error[1].MINUTE"
   IOField "I/O field_12" at 171,119 size 25x19; FormatPattern 999
      ProcessValue <- "Data_DTLData_DTL_Mesin Error[1].HOUR"
   TextField "Text field_8" at 27,119 size 145x19; Text 'Error'
   TextField "Text field_2" at 171,48 size 25x19; Text 'Hour'
   IOField "I/O field_6" at 6,17 size 109x15; FormatPattern 9999999999999999999999999999999999999999
      ProcessValue <- "Data_DTL1_Cur_ShiftA_1"
   TextField "Text field_9" at 120,17 size 18x13; Text 'S/D'
   IOField "I/O field_7" at 143,17 size 109x15; FormatPattern 9999999999999999999999999999999999999999
      ProcessValue <- "Data_DTL1_Cur_ShiftB_1"
   IOField "I/O field_16" at 219,138 size 25x19; FormatPattern 999
      ProcessValue <- "Data_DTLData_Total Time Machine[1].SECOND"
   IOField "I/O field_17" at 195,138 size 25x19; FormatPattern 999
      ProcessValue <- "Data_DTLData_Total Time Machine[1].MINUTE"
   IOField "I/O field_18" at 171,138 size 25x19; FormatPattern 999
      ProcessValue <- "Data_DTLData_Total Time Machine[1].HOUR"
   TextField "Text field_10" at 27,138 size 145x19; Text 'Total'
   IOField "I/O field_27" at 253,16 size 66x17; FormatPattern ????????
      ProcessValue <- "Data_String_sDT_Machine id"

screen "St_Time machine data_2" 320x240
   IOField "I/O field_13" at 243,83 size 56x19; FormatPattern 999.99; Unit   %
      ProcessValue <- "Data_Real_%Mesin Stop[2]"
   IOField "I/O field_14" at 243,101 size 56x19; FormatPattern 999.99; Unit   %
      ProcessValue <- "Data_Real_%Mesin Run Baypass[2]"
   IOField "I/O field_11" at 243,66 size 56x19; FormatPattern 999.99; Unit   %
      ProcessValue <- "Data_Real_%Mesin Run[2]"
   Button "Button_1" at 46,213 size 90x25; TextOff 'Statistic Data'
      on Click: ActivateScreen("St_Data Statistic", 0)
   Button "Button_3" at 1,213 size 41x25; TextOff 'Main Page'; PictureOff "Home"
      on Click: ActivateScreen("Main Page", 0)
   Button "Button_2" at 237,213 size 80x25; TextOff 'Next page -->'; TextOn 'Page 3'
      on Click: ActivateScreen("St_Error Counter_2", 0)
   TextField "Text field_1" at 3,0 size 155x18; Text 'CURRENT SHIFT MINUS 2'
   TextField "Text field_31" at 7,101 size 21x19; Text '3'
   TextField "Text field_30" at 7,83 size 21x19; Text '2'
   TextField "Text field_29" at 7,66 size 21x19; Text '1'
   TextField "Text field_28" at 7,48 size 21x19; Text 'No'
   IOField "I/O field_21" at 219,83 size 25x19; FormatPattern 999
      ProcessValue <- "Data_DTLData_DTL_Mesin Stop[2].SECOND"
   IOField "I/O field_22" at 195,83 size 25x19; FormatPattern 999
      ProcessValue <- "Data_DTLData_DTL_Mesin Stop[2].MINUTE"
   IOField "I/O field_23" at 171,84 size 25x19; FormatPattern 999
      ProcessValue <- "Data_DTLData_DTL_Mesin Stop[2].HOUR"
   TextField "Text field_25" at 27,83 size 145x19; Text 'Stop'
   IOField "I/O field_4" at 219,101 size 25x19; FormatPattern 999
      ProcessValue <- "Data_DTLData_DTL_Mesin Run Baypass[2].SECOND"
   IOField "I/O field_5" at 195,101 size 25x19; FormatPattern 999
      ProcessValue <- "Data_DTLData_DTL_Mesin Run Baypass[2].MINUTE"
   IOField "I/O field_9" at 171,101 size 25x19; FormatPattern 999
      ProcessValue <- "Data_DTLData_DTL_Mesin Run Baypass[2].HOUR"
   TextField "Text field_12" at 219,48 size 25x19; Text 'Sec'
   TextField "Text field_11" at 195,48 size 25x19; Text 'Min'
   IOField "I/O field_2" at 219,66 size 25x19; FormatPattern 999
      ProcessValue <- "Data_DTLData_DTL_Mesin Run[2].SECOND"
   IOField "I/O field_3" at 195,66 size 25x19; FormatPattern 999
      ProcessValue <- "Data_DTLData_DTL_Mesin Run[2].MINUTE"
   TextField "Text field_3" at 27,48 size 145x19; Text 'Time Counter Machine'
   TextField "Text field_4" at 27,66 size 145x19; Text 'Running'
   TextField "Text field_5" at 27,101 size 145x19; Text 'Running Bypass'
   IOField "I/O field_24" at 171,66 size 25x19; FormatPattern 999
      ProcessValue <- "Data_DTLData_DTL_Mesin Run[2].HOUR"
   Button "Button_4" at 151,213 size 80x25; TextOff '<-- Back Page'; TextOn 'Page 1'
      on Click: ActivateScreen("St_Quantity Data_2", 0)
   TextField "Text field_6" at 260,0 size 57x15; Text 'Page 2 of 3'
   IOField "I/O field_1" at 243,119 size 56x19; FormatPattern 999.99; Unit   %
      ProcessValue <- "Data_Real_%Mesin Error[2]"
   TextField "Text field_7" at 7,119 size 21x19; Text '4'
   IOField "I/O field_8" at 219,119 size 25x19; FormatPattern 999
      ProcessValue <- "Data_DTLData_DTL_Mesin Error[2].SECOND"
   IOField "I/O field_10" at 195,119 size 25x19; FormatPattern 999
      ProcessValue <- "Data_DTLData_DTL_Mesin Error[2].MINUTE"
   IOField "I/O field_12" at 171,119 size 25x19; FormatPattern 999
      ProcessValue <- "Data_DTLData_DTL_Mesin Error[2].HOUR"
   TextField "Text field_8" at 27,119 size 145x19; Text 'Error'
   TextField "Text field_2" at 171,48 size 25x19; Text 'Hour'
   IOField "I/O field_6" at 6,17 size 109x15; FormatPattern 9999999999999999999999999999999999999999
      ProcessValue <- "Data_DTL1_Cur_ShiftA_2"
   TextField "Text field_9" at 120,17 size 18x13; Text 'S/D'
   IOField "I/O field_7" at 143,17 size 109x15; FormatPattern 9999999999999999999999999999999999999999
      ProcessValue <- "Data_DTL1_Cur_ShiftB_2"
   IOField "I/O field_16" at 219,138 size 25x19; FormatPattern 999
      ProcessValue <- "Data_DTLData_Total Time Machine[2].SECOND"
   IOField "I/O field_17" at 195,138 size 25x19; FormatPattern 999
      ProcessValue <- "Data_DTLData_Total Time Machine[2].MINUTE"
   IOField "I/O field_18" at 171,138 size 25x19; FormatPattern 999
      ProcessValue <- "Data_DTLData_Total Time Machine[2].HOUR"
   TextField "Text field_10" at 27,138 size 145x19; Text 'Total'
   IOField "I/O field_27" at 253,16 size 66x17; FormatPattern ????????
      ProcessValue <- "Data_String_sDT_Machine id"

screen "St_Time machine data_3" 320x240
   IOField "I/O field_13" at 243,83 size 56x19; FormatPattern 999.99; Unit   %
      ProcessValue <- "Data_Real_%Mesin Stop[3]"
   IOField "I/O field_14" at 243,101 size 56x19; FormatPattern 999.99; Unit   %
      ProcessValue <- "Data_Real_%Mesin Run Baypass[3]"
   IOField "I/O field_11" at 243,66 size 56x19; FormatPattern 999.99; Unit   %
      ProcessValue <- "Data_Real_%Mesin Run[3]"
   Button "Button_1" at 46,213 size 90x25; TextOff 'Statistic Data'
      on Click: ActivateScreen("St_Data Statistic", 0)
   Button "Button_3" at 1,213 size 41x25; TextOff 'Main Page'; PictureOff "Home"
      on Click: ActivateScreen("Main Page", 0)
   Button "Button_2" at 237,213 size 80x25; TextOff 'Next page -->'; TextOn 'Page 3'
      on Click: ActivateScreen("St_Error Counter_3", 0)
   TextField "Text field_1" at 3,0 size 155x18; Text 'CURRENT SHIFT MINUS 3'
   TextField "Text field_31" at 7,101 size 21x19; Text '3'
   TextField "Text field_30" at 7,83 size 21x19; Text '2'
   TextField "Text field_29" at 7,66 size 21x19; Text '1'
   TextField "Text field_28" at 7,48 size 21x19; Text 'No'
   IOField "I/O field_21" at 219,83 size 25x19; FormatPattern 999
      ProcessValue <- "Data_DTLData_DTL_Mesin Stop[3].SECOND"
   IOField "I/O field_22" at 195,83 size 25x19; FormatPattern 999
      ProcessValue <- "Data_DTLData_DTL_Mesin Stop[3].MINUTE"
   IOField "I/O field_23" at 171,84 size 25x19; FormatPattern 999
      ProcessValue <- "Data_DTLData_DTL_Mesin Stop[3].HOUR"
   TextField "Text field_25" at 27,83 size 145x19; Text 'Stop'
   IOField "I/O field_4" at 219,101 size 25x19; FormatPattern 999
      ProcessValue <- "Data_DTLData_DTL_Mesin Run Baypass[3].SECOND"
   IOField "I/O field_5" at 195,101 size 25x19; FormatPattern 999
      ProcessValue <- "Data_DTLData_DTL_Mesin Run Baypass[3].MINUTE"
   IOField "I/O field_9" at 171,101 size 25x19; FormatPattern 999
      ProcessValue <- "Data_DTLData_DTL_Mesin Run Baypass[3].HOUR"
   TextField "Text field_12" at 219,48 size 25x19; Text 'Sec'
   TextField "Text field_11" at 195,48 size 25x19; Text 'Min'
   IOField "I/O field_2" at 219,66 size 25x19; FormatPattern 999
      ProcessValue <- "Data_DTLData_DTL_Mesin Run[3].SECOND"
   IOField "I/O field_3" at 195,66 size 25x19; FormatPattern 999
      ProcessValue <- "Data_DTLData_DTL_Mesin Run[3].MINUTE"
   TextField "Text field_3" at 27,48 size 145x19; Text 'Time Counter Machine'
   TextField "Text field_4" at 27,66 size 145x19; Text 'Running'
   TextField "Text field_5" at 27,101 size 145x19; Text 'Running Bypass'
   IOField "I/O field_24" at 171,66 size 25x19; FormatPattern 999
      ProcessValue <- "Data_DTLData_DTL_Mesin Run[3].HOUR"
   Button "Button_4" at 151,213 size 80x25; TextOff '<-- Back Page'; TextOn 'Page 1'
      on Click: ActivateScreen("St_Quantity Data_3", 0)
   TextField "Text field_6" at 260,0 size 57x15; Text 'Page 2 of 3'
   IOField "I/O field_1" at 243,119 size 56x19; FormatPattern 999.99; Unit   %
      ProcessValue <- "Data_Real_%Mesin Error[3]"
   TextField "Text field_7" at 7,119 size 21x19; Text '4'
   IOField "I/O field_8" at 219,119 size 25x19; FormatPattern 999
      ProcessValue <- "Data_DTLData_DTL_Mesin Error[3].SECOND"
   IOField "I/O field_10" at 195,119 size 25x19; FormatPattern 999
      ProcessValue <- "Data_DTLData_DTL_Mesin Error[3].MINUTE"
   IOField "I/O field_12" at 171,119 size 25x19; FormatPattern 999
      ProcessValue <- "Data_DTLData_DTL_Mesin Error[3].HOUR"
   TextField "Text field_8" at 27,119 size 145x19; Text 'Error'
   TextField "Text field_2" at 171,48 size 25x19; Text 'Hour'
   IOField "I/O field_6" at 6,17 size 109x15; FormatPattern 9999999999999999999999999999999999999999
      ProcessValue <- "Data_DTL1_Cur_ShiftA_3"
   TextField "Text field_9" at 120,17 size 18x13; Text 'S/D'
   IOField "I/O field_7" at 143,17 size 109x15; FormatPattern 9999999999999999999999999999999999999999
      ProcessValue <- "Data_DTL1_Cur_ShiftB_3"
   IOField "I/O field_16" at 219,138 size 25x19; FormatPattern 999
      ProcessValue <- "Data_DTLData_Total Time Machine[3].SECOND"
   IOField "I/O field_17" at 195,138 size 25x19; FormatPattern 999
      ProcessValue <- "Data_DTLData_Total Time Machine[3].MINUTE"
   IOField "I/O field_18" at 171,138 size 25x19; FormatPattern 999
      ProcessValue <- "Data_DTLData_Total Time Machine[3].HOUR"
   TextField "Text field_10" at 27,138 size 145x19; Text 'Total'
   IOField "I/O field_27" at 253,16 size 66x17; FormatPattern ????????
      ProcessValue <- "Data_String_sDT_Machine id"

